(* Logix 5000 project; controller PLC_MCC1300_75F1 vendor 1 type 14 code 166 rev 32.11; software revision 32.04; part 54 of 83 *)
(* tags used below, declared in another part *)
   AUX_tConvoy_SL_NULL : UDT_Convoy_SL;
   CONST_dDest_Cullet : DINT;
   CONST_dDest_Stk : DINT;
   CONST_rgdDestMask : DINT[32];   // Destination Mask
   CONST_tPlant : UDT_PLANT_CONSTANTS;
   GP_CheckIdPlatePresent : GP_CheckIdPlatePresent;
   GP_RampSpace : GP_RampSpace;
   Gp_SpaceConvUtilities_V1 : GP_SpaceConvUtilities_V1;
   GP_TrackingSearchPlate : GP_TrackingSearchPlate;
   M310B_SpaceConv_Utilities : SpaceConv_Utilities;
   M310Popup : MAC_Popup_ZC[2];
   M310Popup_HMW : MAC_Popup_ZC_HMW[2];
   M310Popup_SL_DATA : UDT_Convoy_SL;
   M310Popup_tSearchPlateChangeFromCS4401 : GP_TrackingSearchPlate_STC;
   M310Popup_xDrivePosEnable : BOOL;
   M310Popup_xEndRiseWaitingForCondition : BOOL;
   M311 : MAC_Conveyor;
   M311_ALM : MAC_Conveyor_ALM;
   M311_Data : UDT_Convoy_SL;
   M311_HMW : MAC_Conveyor_HMW;
   M311_SpaceConv_Utilities : SpaceConv_Utilities;
   M311_xPlateCullet : BOOL;
   M311A : MAC_Rotator;
   M311A_HMW : MAC_Rotator_HMW;
   M312 : MAC_Conveyor_Single;
   M312_SpaceConv_Utilities : SpaceConv_Utilities;
   M350Popup : MAC_Popup_ZC;
   TMP_d : DINT;
   TMP_dConveyorNumberForZoneCleaning : DINT;
   TMP_dIndexCap : DINT;
   TMP_dMaskAllowed : DINT;
   TMP_dOffsetLoadUnload_cmm : DINT;
   TMP_dPhEndPosition_cmm : DINT;
   TMP_dStartSearch : DINT;
   TMP_dStopSearch : DINT;
   TMP_rgxId : DINT[10];
   TMP_xAllLiteToCullet : BOOL;
   TMP_xAtLeastOneForSideLeg : BOOL;
   TMP_xConveyorInvolvedInCleaning : BOOL;
   TMP_xConveyorOfStartCleaning : BOOL;
   TMP_xCulletPresent : BOOL;
   TMP_xDummy : BOOL;
   TMP_xEnableLoadUnload : BOOL;
   TMP_xEnableZoneCleaning : BOOL;
   TMP_xLiteThisDestPresent : BOOL;
   xAlwaysOFF : BOOL;
   xAlwaysON : BOOL;
   Z300_BufferPlate : UDT_LINE_BUFFER_PLATE;
   Z300_Conveyor : UDT_StandConv[29];
   Z300_LineTracking : UDT_LINE_TRACKING;
   Z301 : MAC_Zone_ML;
   Z401 : MAC_Zone;
   Z401_HMR : MAC_Zone_HMR;
   Z401_HMW : MAC_Zone_HMW;
(* MainProgram, continued *)

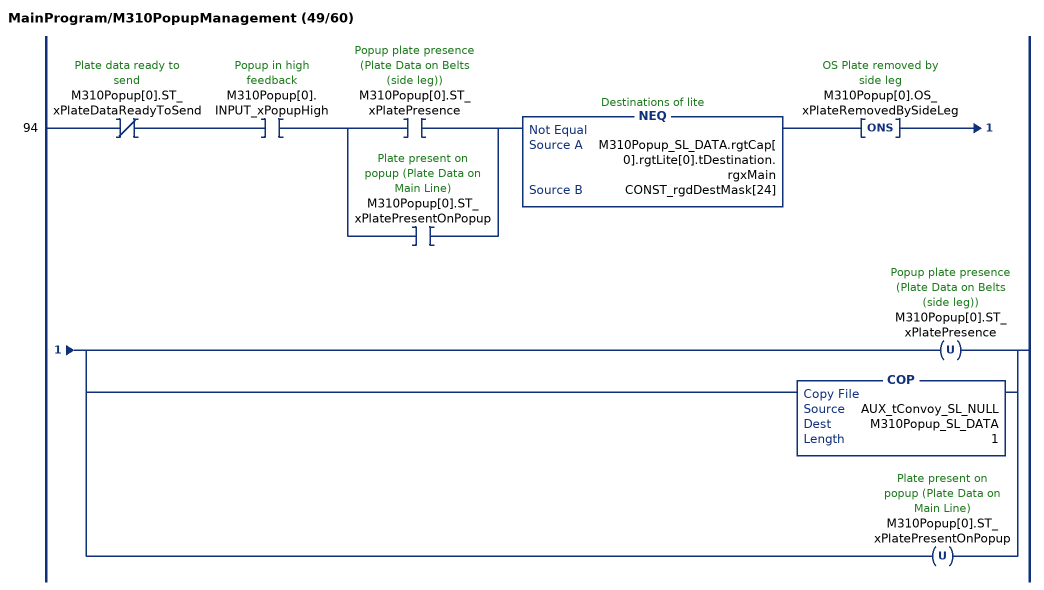
   [picture p865: MainProgram/M310PopupManagement rungs 94-94]
   94: XIO(M310Popup[0].ST_xPlateDataReadyToSend)XIC(M310Popup[0].INPUT_xPopupHigh)[XIC(M310Popup[0].ST_xPlatePresence) ,XIC(M310Popup[0].ST_xPlatePresentOnPopup) ]NEQ(M310Popup_SL_DATA.rgtCap[0].rgtLite[0].tDestination.rgxMain,CONST_rgdDestMask[24])ONS(M310Popup[0].OS_xPlateRemovedBySideLeg)[OTU(M310Popup[0].ST_xPlatePresence) ,COP(AUX_tConvoy_SL_NULL,M310Popup_SL_DATA,1) ,OTU(M310Popup[0].ST_xPlatePresentOnPopup) ];
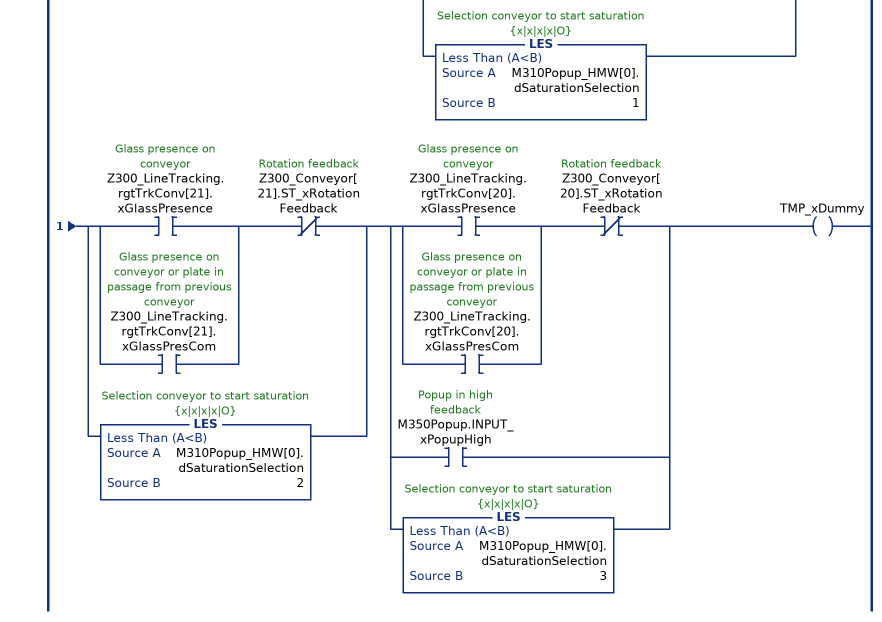
   // #####_SATURATION_#####
   95: GRT(M310Popup_HMW[0].dSaturationSelection,0)XIC(Z301.ST_xCycleON)[[[XIC(Z300_LineTracking.rgtTrkConv[22].xGlassPresence) ,XIC(Z300_LineTracking.rgtTrkConv[23].xGlassPresence) ,XIC(Z300_LineTracking.rgtTrkConv[24].xGlassPresence) ,XIC(Z300_LineTracking.rgtTrkConv[22].xGlassPresCom) ,XIC(Z300_LineTracking.rgtTrkConv[23].xGlassPresCom) ,XIC(Z300_LineTracking.rgtTrkConv[24].xGlassPresCom) ] [XIO(Z300_Conveyor[22].ST_xRotationFeedback) ,XIO(Z300_Conveyor[23].ST_xRotationFeedback) ,XIO(Z300_Conveyor[24].ST_xRotationFeedback) ] ,XIO(xAlwaysOFF) [XIC(M310Popup[0].ST_xPlatePresence) XIC(M310Popup[0].INPUT_xPopupHigh) ,[XIO(M310Popup[0].ST_xInitialConditionForRise) ,XIO(M310Popup[1].ST_xInitialConditionForRise) ] ] ] ,LES(M310Popup_HMW[0].dSaturationSelection,1) ][[XIC(Z300_LineTracking.rgtTrkConv[21].xGlassPresence) ,XIC(Z300_LineTracking.rgtTrkConv[21].xGlassPresCom) ] XIO(Z300_Conveyor[21].ST_xRotationFeedback) ,LES(M310Popup_HMW[0].dSaturationSelection,2) ][[[XIC(Z300_LineTracking.rgtTrkConv[20].xGlassPresence) ,XIC(Z300_LineTracking.rgtTrkConv[20].xGlassPresCom) ] XIO(Z300_Conveyor[20].ST_xRotationFeedback) ,XIC(M350Popup.INPUT_xPopupHigh) ] ,LES(M310Popup_HMW[0].dSaturationSelection,3) ]OTE(TMP_xDummy);
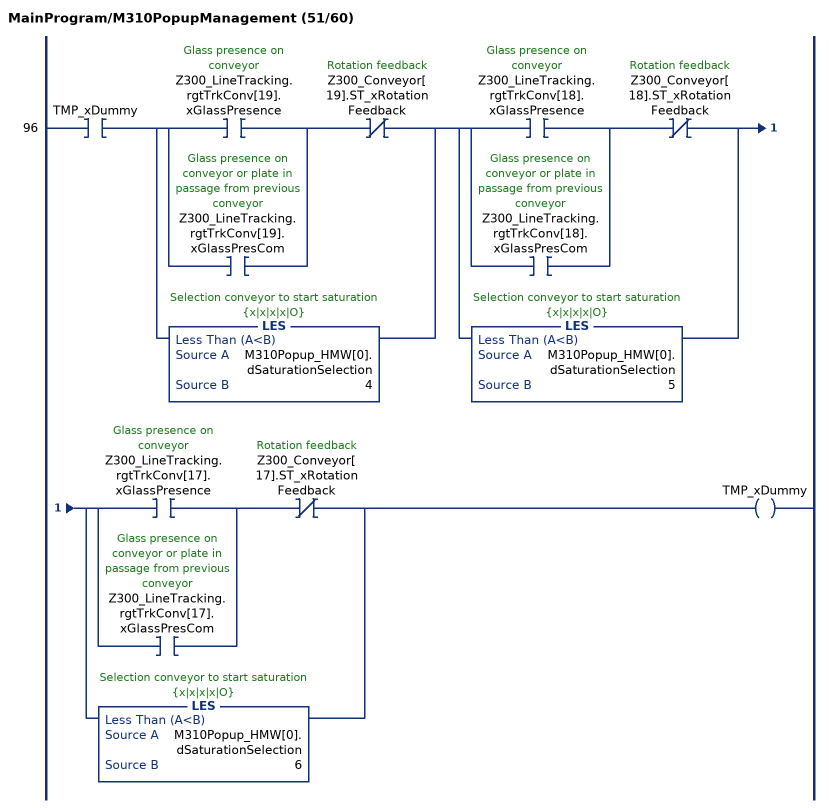
   96: XIC(TMP_xDummy)[[XIC(Z300_LineTracking.rgtTrkConv[19].xGlassPresence) ,XIC(Z300_LineTracking.rgtTrkConv[19].xGlassPresCom) ] XIO(Z300_Conveyor[19].ST_xRotationFeedback) ,LES(M310Popup_HMW[0].dSaturationSelection,4) ][[XIC(Z300_LineTracking.rgtTrkConv[18].xGlassPresence) ,XIC(Z300_LineTracking.rgtTrkConv[18].xGlassPresCom) ] XIO(Z300_Conveyor[18].ST_xRotationFeedback) ,LES(M310Popup_HMW[0].dSaturationSelection,5) ][[XIC(Z300_LineTracking.rgtTrkConv[17].xGlassPresence) ,XIC(Z300_LineTracking.rgtTrkConv[17].xGlassPresCom) ] XIO(Z300_Conveyor[17].ST_xRotationFeedback) ,LES(M310Popup_HMW[0].dSaturationSelection,6) ]OTE(TMP_xDummy);
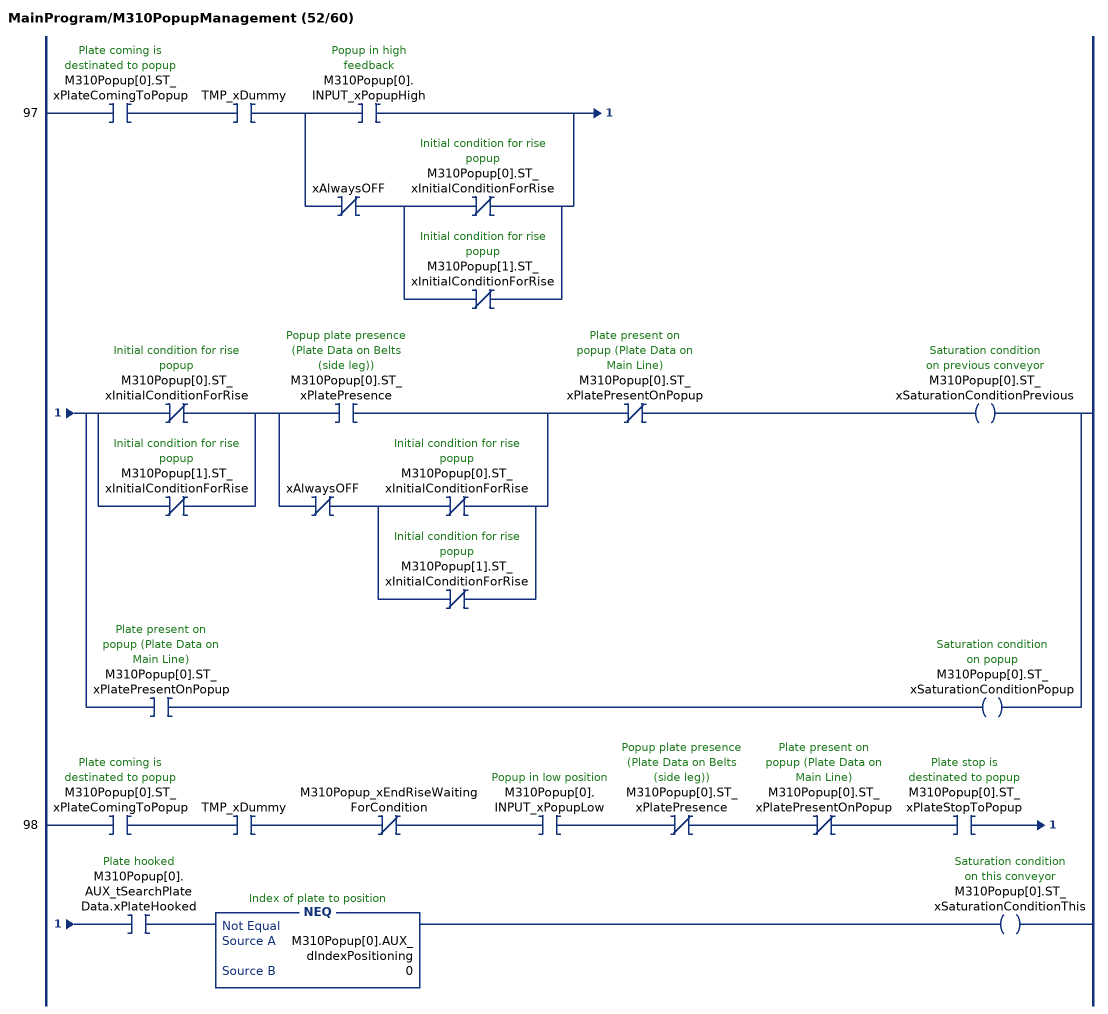
   97: XIC(M310Popup[0].ST_xPlateComingToPopup)XIC(TMP_xDummy)[XIC(M310Popup[0].INPUT_xPopupHigh) ,XIO(xAlwaysOFF) [XIO(M310Popup[0].ST_xInitialConditionForRise) ,XIO(M310Popup[1].ST_xInitialConditionForRise) ] ][[XIO(M310Popup[0].ST_xInitialConditionForRise) ,XIO(M310Popup[1].ST_xInitialConditionForRise) ] [XIC(M310Popup[0].ST_xPlatePresence) ,XIO(xAlwaysOFF) [XIO(M310Popup[0].ST_xInitialConditionForRise) ,XIO(M310Popup[1].ST_xInitialConditionForRise) ] ] XIO(M310Popup[0].ST_xPlatePresentOnPopup) OTE(M310Popup[0].ST_xSaturationConditionPrevious) ,XIC(M310Popup[0].ST_xPlatePresentOnPopup) OTE(M310Popup[0].ST_xSaturationConditionPopup) ];
   98: XIC(M310Popup[0].ST_xPlateComingToPopup)XIC(TMP_xDummy)XIO(M310Popup_xEndRiseWaitingForCondition)XIC(M310Popup[0].INPUT_xPopupLow)XIO(M310Popup[0].ST_xPlatePresence)XIO(M310Popup[0].ST_xPlatePresentOnPopup)XIC(M310Popup[0].ST_xPlateStopToPopup)XIC(M310Popup[0].AUX_tSearchPlateData.xPlateHooked)NEQ(M310Popup[0].AUX_dIndexPositioning,0)OTE(M310Popup[0].ST_xSaturationConditionThis);
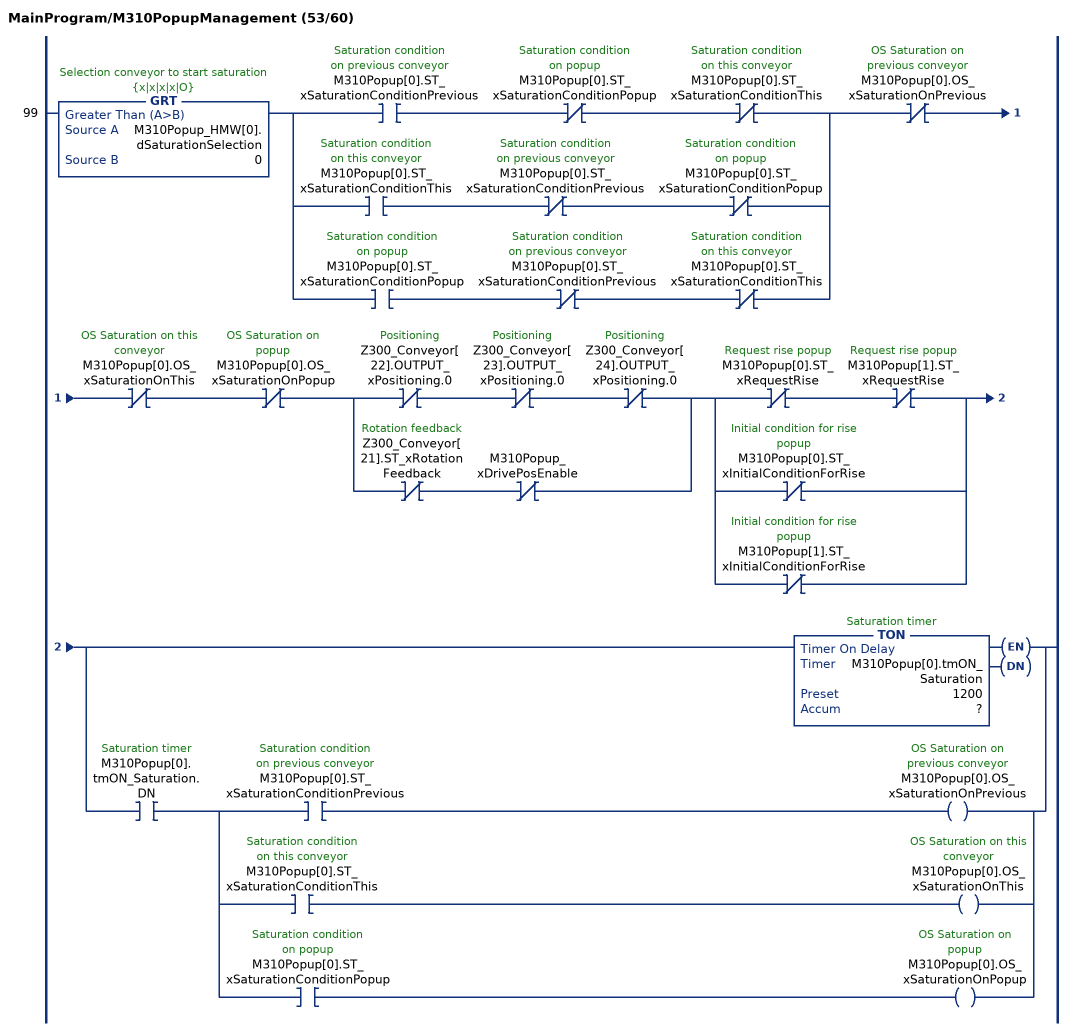
   99: GRT(M310Popup_HMW[0].dSaturationSelection,0)[XIC(M310Popup[0].ST_xSaturationConditionPrevious) XIO(M310Popup[0].ST_xSaturationConditionPopup) XIO(M310Popup[0].ST_xSaturationConditionThis) ,XIC(M310Popup[0].ST_xSaturationConditionThis) XIO(M310Popup[0].ST_xSaturationConditionPrevious) XIO(M310Popup[0].ST_xSaturationConditionPopup) ,XIC(M310Popup[0].ST_xSaturationConditionPopup) XIO(M310Popup[0].ST_xSaturationConditionPrevious) XIO(M310Popup[0].ST_xSaturationConditionThis) ]XIO(M310Popup[0].OS_xSaturationOnPrevious)XIO(M310Popup[0].OS_xSaturationOnThis)XIO(M310Popup[0].OS_xSaturationOnPopup)[XIO(Z300_Conveyor[22].OUTPUT_xPositioning.0) XIO(Z300_Conveyor[23].OUTPUT_xPositioning.0) XIO(Z300_Conveyor[24].OUTPUT_xPositioning.0) ,XIO(Z300_Conveyor[21].ST_xRotationFeedback) XIO(M310Popup_xDrivePosEnable) ][XIO(M310Popup[0].ST_xRequestRise) XIO(M310Popup[1].ST_xRequestRise) ,XIO(M310Popup[0].ST_xInitialConditionForRise) ,XIO(M310Popup[1].ST_xInitialConditionForRise) ][TON(M310Popup[0].tmON_Saturation,?,?) ,XIC(M310Popup[0].tmON_Saturation.DN) [XIC(M310Popup[0].ST_xSaturationConditionPrevious) OTE(M310Popup[0].OS_xSaturationOnPrevious) ,XIC(M310Popup[0].ST_xSaturationConditionThis) OTE(M310Popup[0].OS_xSaturationOnThis) ,XIC(M310Popup[0].ST_xSaturationConditionPopup) OTE(M310Popup[0].OS_xSaturationOnPopup) ] ];
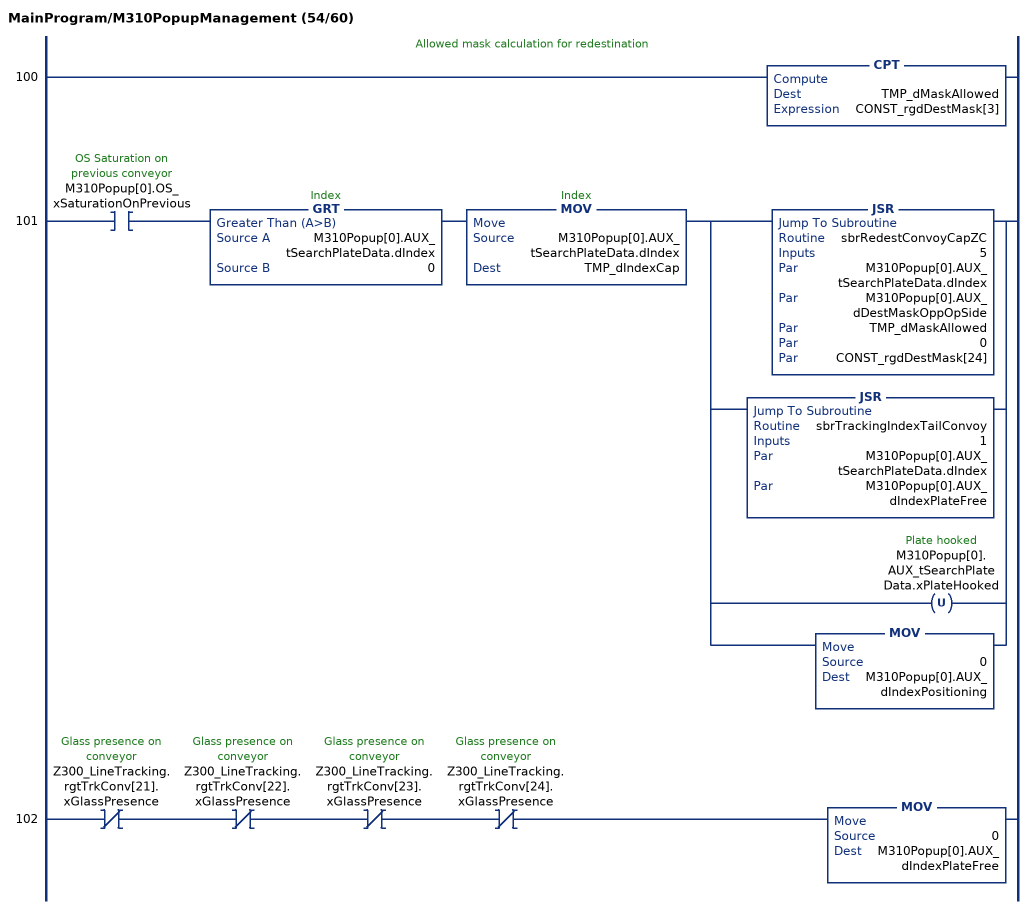
   // Allowed mask calculation for redestination
   100: CPT(TMP_dMaskAllowed,CONST_rgdDestMask[3]);
   101: XIC(M310Popup[0].OS_xSaturationOnPrevious)GRT(M310Popup[0].AUX_tSearchPlateData.dIndex,0)MOV(M310Popup[0].AUX_tSearchPlateData.dIndex,TMP_dIndexCap)[JSR(sbrRedestConvoyCapZC,5,M310Popup[0].AUX_tSearchPlateData.dIndex,M310Popup[0].AUX_dDestMaskOppOpSide,TMP_dMaskAllowed,0,CONST_rgdDestMask[24]) ,JSR(sbrTrackingIndexTailConvoy,1,M310Popup[0].AUX_tSearchPlateData.dIndex,M310Popup[0].AUX_dIndexPlateFree) ,[OTU(M310Popup[0].AUX_tSearchPlateData.xPlateHooked) ,MOV(0,M310Popup[0].AUX_dIndexPositioning) ] ];
   102: XIO(Z300_LineTracking.rgtTrkConv[21].xGlassPresence)XIO(Z300_LineTracking.rgtTrkConv[22].xGlassPresence)XIO(Z300_LineTracking.rgtTrkConv[23].xGlassPresence)XIO(Z300_LineTracking.rgtTrkConv[24].xGlassPresence)MOV(0,M310Popup[0].AUX_dIndexPlateFree);
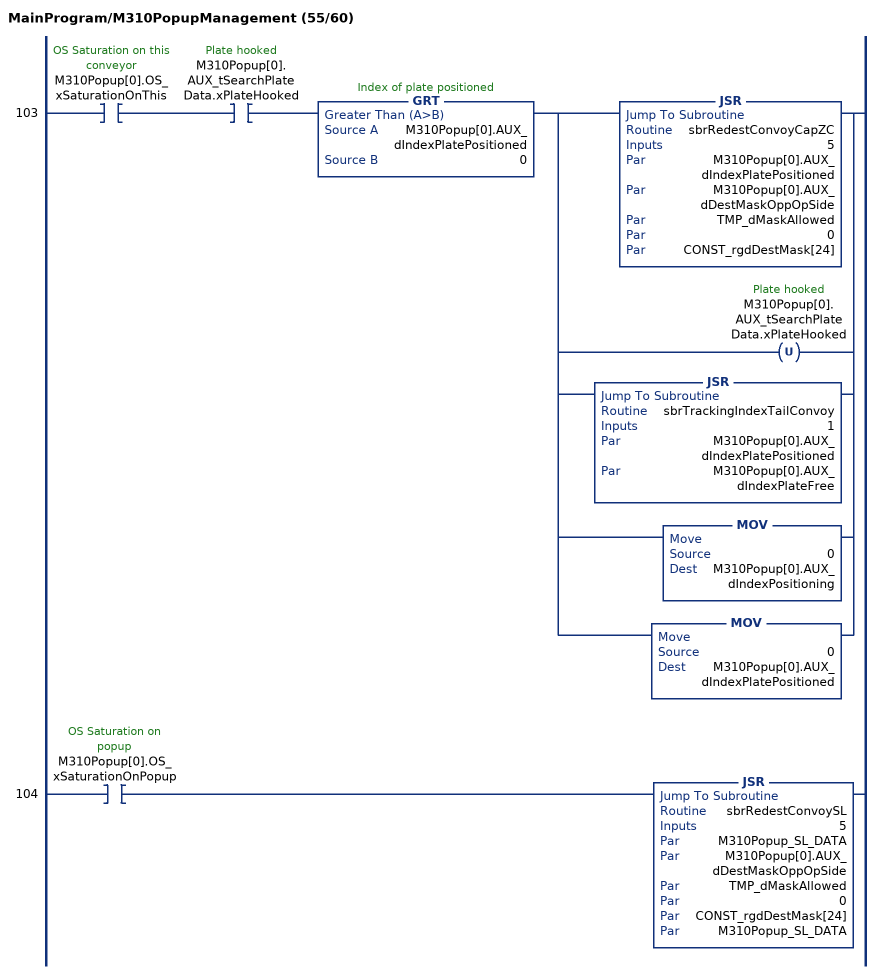
   103: XIC(M310Popup[0].OS_xSaturationOnThis)XIC(M310Popup[0].AUX_tSearchPlateData.xPlateHooked)GRT(M310Popup[0].AUX_dIndexPlatePositioned,0)[JSR(sbrRedestConvoyCapZC,5,M310Popup[0].AUX_dIndexPlatePositioned,M310Popup[0].AUX_dDestMaskOppOpSide,TMP_dMaskAllowed,0,CONST_rgdDestMask[24]) ,OTU(M310Popup[0].AUX_tSearchPlateData.xPlateHooked) ,JSR(sbrTrackingIndexTailConvoy,1,M310Popup[0].AUX_dIndexPlatePositioned,M310Popup[0].AUX_dIndexPlateFree) ,MOV(0,M310Popup[0].AUX_dIndexPositioning) ,MOV(0,M310Popup[0].AUX_dIndexPlatePositioned) ];
   104: XIC(M310Popup[0].OS_xSaturationOnPopup)JSR(sbrRedestConvoySL,5,M310Popup_SL_DATA,M310Popup[0].AUX_dDestMaskOppOpSide,TMP_dMaskAllowed,0,CONST_rgdDestMask[24],M310Popup_SL_DATA);
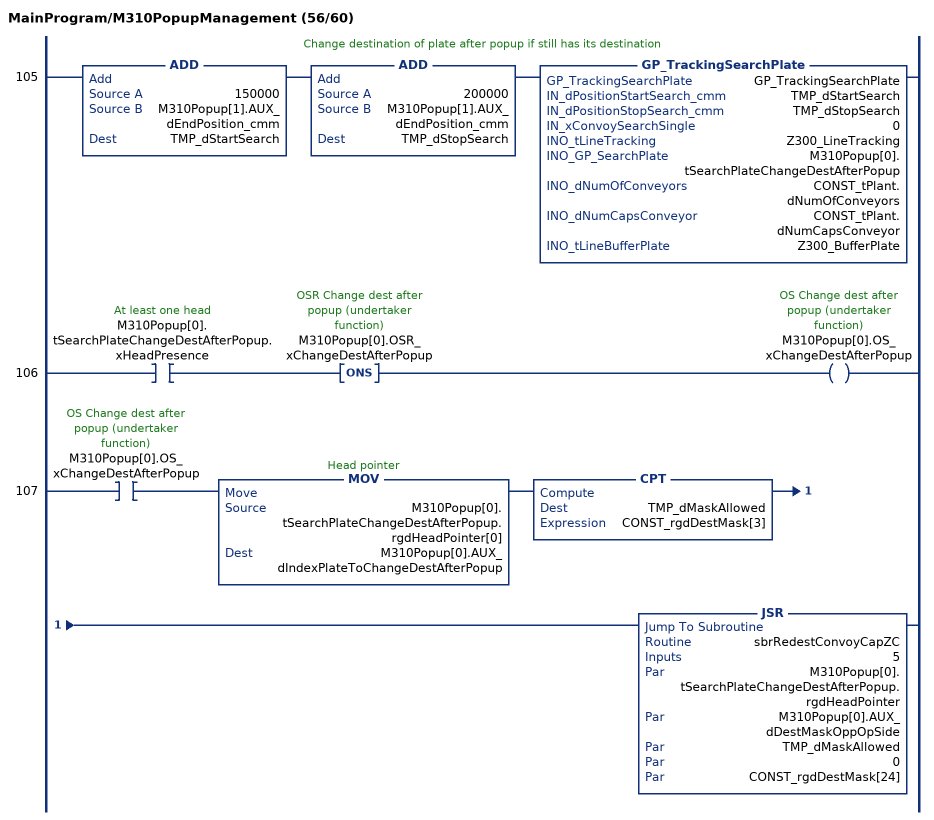
   // Change destination of plate after popup if still has its destination
   105: ADD(150000,M310Popup[1].AUX_dEndPosition_cmm,TMP_dStartSearch)ADD(200000,M310Popup[1].AUX_dEndPosition_cmm,TMP_dStopSearch)GP_TrackingSearchPlate(GP_TrackingSearchPlate,TMP_dStartSearch,TMP_dStopSearch,0,Z300_LineTracking,M310Popup[0].tSearchPlateChangeDestAfterPopup,CONST_tPlant.dNumOfConveyors,CONST_tPlant.dNumCapsConveyor,Z300_BufferPlate);
   106: XIC(M310Popup[0].tSearchPlateChangeDestAfterPopup.xHeadPresence)ONS(M310Popup[0].OSR_xChangeDestAfterPopup)OTE(M310Popup[0].OS_xChangeDestAfterPopup);
   107: XIC(M310Popup[0].OS_xChangeDestAfterPopup)MOV(M310Popup[0].tSearchPlateChangeDestAfterPopup.rgdHeadPointer[0],M310Popup[0].AUX_dIndexPlateToChangeDestAfterPopup)CPT(TMP_dMaskAllowed,CONST_rgdDestMask[3])JSR(sbrRedestConvoyCapZC,5,M310Popup[0].tSearchPlateChangeDestAfterPopup.rgdHeadPointer,M310Popup[0].AUX_dDestMaskOppOpSide,TMP_dMaskAllowed,0,CONST_rgdDestMask[24]);
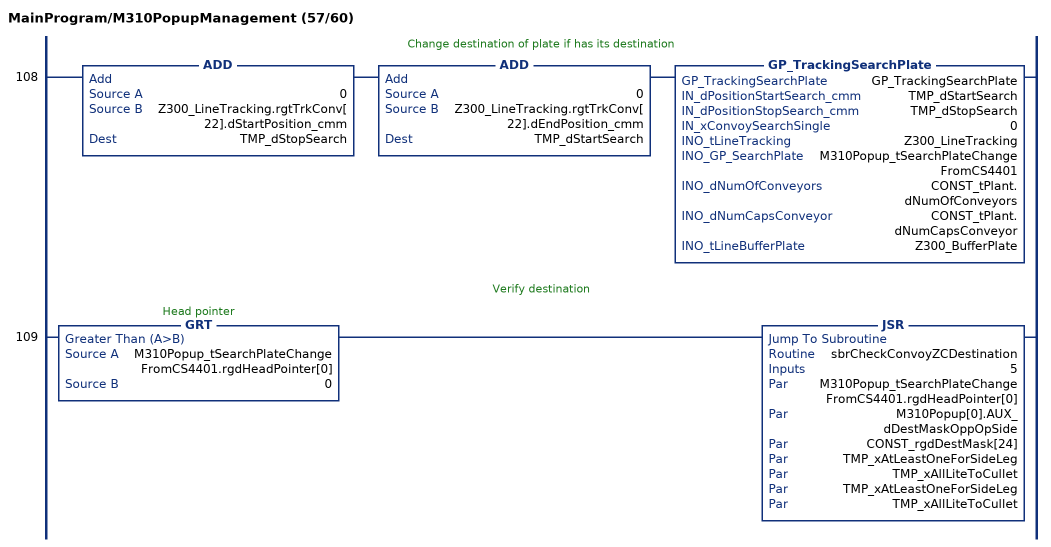
   // Change destination of plate if has its destination
   108: ADD(0,Z300_LineTracking.rgtTrkConv[22].dStartPosition_cmm,TMP_dStopSearch)ADD(0,Z300_LineTracking.rgtTrkConv[22].dEndPosition_cmm,TMP_dStartSearch)GP_TrackingSearchPlate(GP_TrackingSearchPlate,TMP_dStartSearch,TMP_dStopSearch,0,Z300_LineTracking,M310Popup_tSearchPlateChangeFromCS4401,CONST_tPlant.dNumOfConveyors,CONST_tPlant.dNumCapsConveyor,Z300_BufferPlate);
   // Verify destination
   109: GRT(M310Popup_tSearchPlateChangeFromCS4401.rgdHeadPointer[0],0)JSR(sbrCheckConvoyZCDestination,5,M310Popup_tSearchPlateChangeFromCS4401.rgdHeadPointer[0],M310Popup[0].AUX_dDestMaskOppOpSide,CONST_rgdDestMask[24],TMP_xAtLeastOneForSideLeg,TMP_xAllLiteToCullet,TMP_xAtLeastOneForSideLeg,TMP_xAllLiteToCullet);
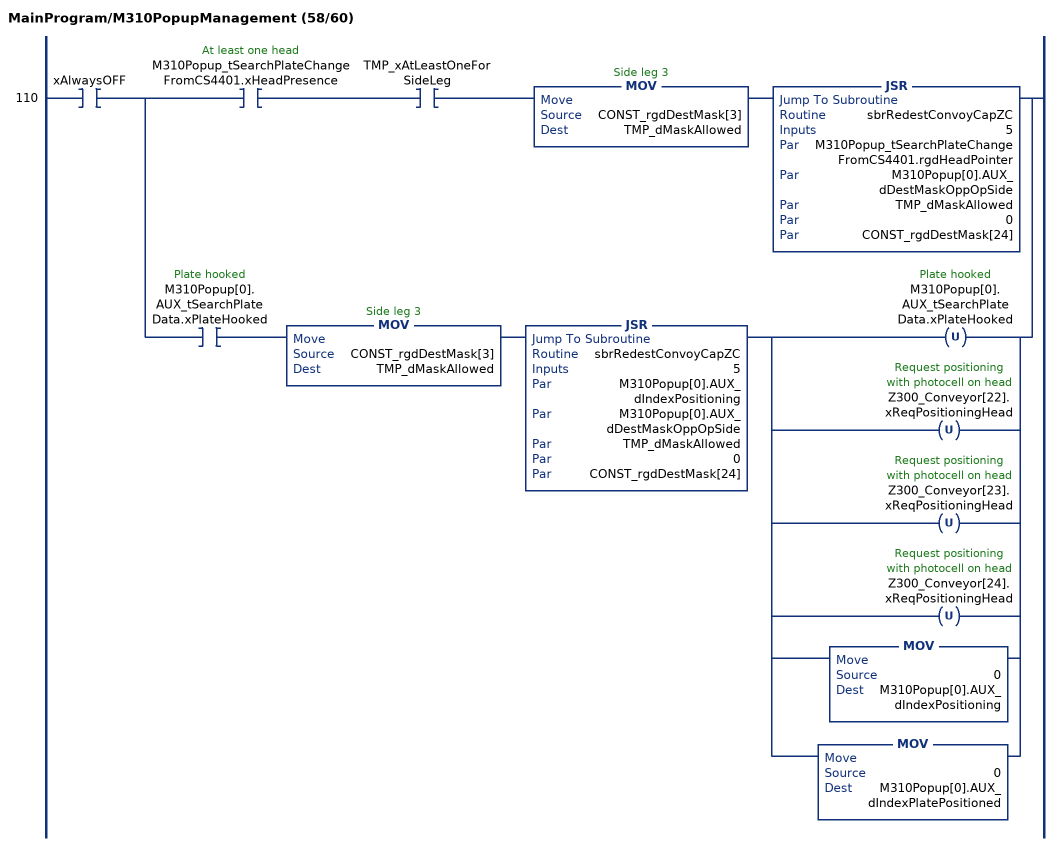
   110: XIC(xAlwaysOFF)[XIC(M310Popup_tSearchPlateChangeFromCS4401.xHeadPresence) XIC(TMP_xAtLeastOneForSideLeg) MOV(CONST_rgdDestMask[3],TMP_dMaskAllowed) JSR(sbrRedestConvoyCapZC,5,M310Popup_tSearchPlateChangeFromCS4401.rgdHeadPointer,M310Popup[0].AUX_dDestMaskOppOpSide,TMP_dMaskAllowed,0,CONST_rgdDestMask[24]) ,XIC(M310Popup[0].AUX_tSearchPlateData.xPlateHooked) MOV(CONST_rgdDestMask[3],TMP_dMaskAllowed) JSR(sbrRedestConvoyCapZC,5,M310Popup[0].AUX_dIndexPositioning,M310Popup[0].AUX_dDestMaskOppOpSide,TMP_dMaskAllowed,0,CONST_rgdDestMask[24]) [OTU(M310Popup[0].AUX_tSearchPlateData.xPlateHooked) ,OTU(Z300_Conveyor[22].xReqPositioningHead) ,OTU(Z300_Conveyor[23].xReqPositioningHead) ,OTU(Z300_Conveyor[24].xReqPositioningHead) ,MOV(0,M310Popup[0].AUX_dIndexPositioning) ,MOV(0,M310Popup[0].AUX_dIndexPlatePositioned) ] ];
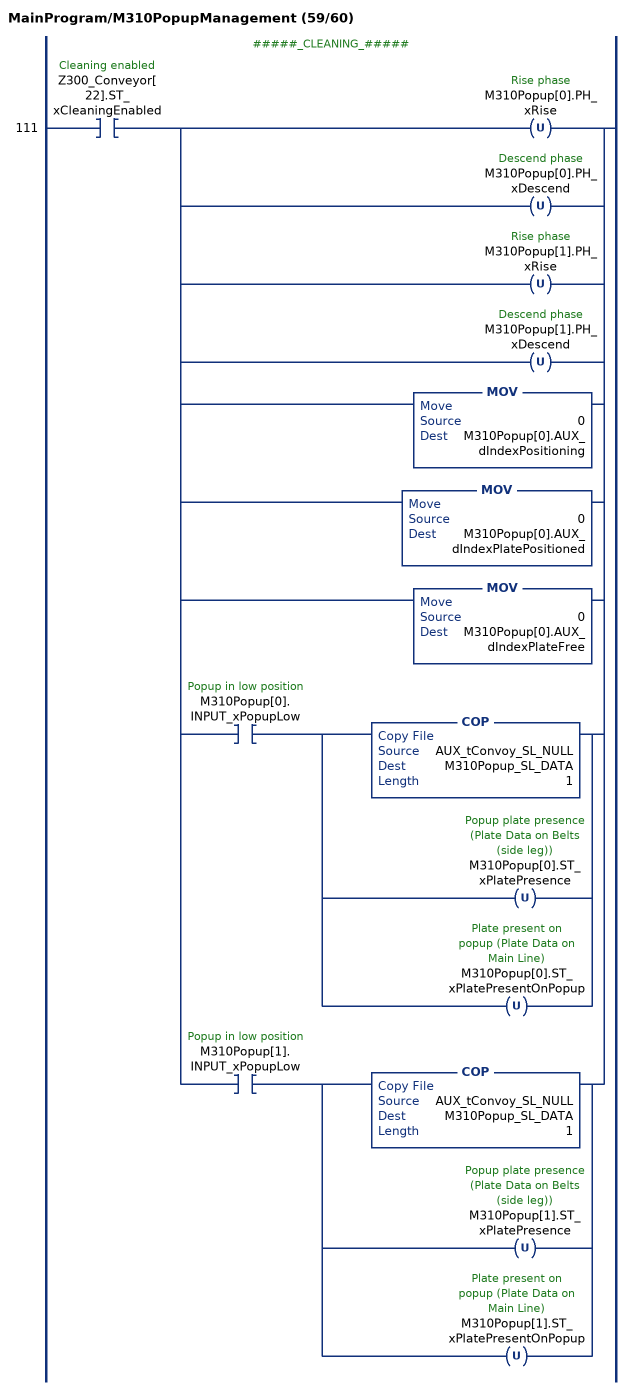
   // #####_CLEANING_#####
   111: XIC(Z300_Conveyor[22].ST_xCleaningEnabled)[OTU(M310Popup[0].PH_xRise) ,OTU(M310Popup[0].PH_xDescend) ,OTU(M310Popup[1].PH_xRise) ,OTU(M310Popup[1].PH_xDescend) ,MOV(0,M310Popup[0].AUX_dIndexPositioning) ,MOV(0,M310Popup[0].AUX_dIndexPlatePositioned) ,MOV(0,M310Popup[0].AUX_dIndexPlateFree) ,XIC(M310Popup[0].INPUT_xPopupLow) [COP(AUX_tConvoy_SL_NULL,M310Popup_SL_DATA,1) ,OTU(M310Popup[0].ST_xPlatePresence) ,OTU(M310Popup[0].ST_xPlatePresentOnPopup) ] ,XIC(M310Popup[1].INPUT_xPopupLow) [COP(AUX_tConvoy_SL_NULL,M310Popup_SL_DATA,1) ,OTU(M310Popup[1].ST_xPlatePresence) ,OTU(M310Popup[1].ST_xPlatePresentOnPopup) ] ];